   "86_Times_STEP_MAX_TIME_STP_540" : Time = PLC "86_Times".STEP_MAX_TIME_STP_540, 1 s
   "86_Times_STEP_MAX_TIME_STP_550" : Time = PLC "86_Times".STEP_MAX_TIME_STP_550, 1 s
   "86_Times_STEP_MAX_TIME_STP_560" : Time = PLC "86_Times".STEP_MAX_TIME_STP_560, 1 s
   "86_Times_STEP_MAX_TIME_STP_570" : Time = PLC "86_Times".STEP_MAX_TIME_STP_570, 1 s
   "86_Times_STEP_MAX_TIME_STP_580" : Time = PLC "86_Times".STEP_MAX_TIME_STP_580, 1 s
   "86_Times_STEP_MAX_TIME_STP_590" : Time = PLC "86_Times".STEP_MAX_TIME_STP_590, 1 s
   "86_Times_STEP_MAX_TIME_STP_600" : Time = PLC "86_Times".STEP_MAX_TIME_STP_600, 1 s
   "86_Times_STEP_MAX_TIME_STP_610" : Time = PLC "86_Times".STEP_MAX_TIME_STP_610, 1 s
   "86_Times_STEP_MAX_TIME_STP_620" : Time = PLC "86_Times".STEP_MAX_TIME_STP_620, 1 s
   "86_Times_STEP_MAX_TIME_STP_630" : Time = PLC "86_Times".STEP_MAX_TIME_STP_630, 1 s
   "150_GCU_LCL_CNTRL_DB_LCL_CNTRL_ACTV" : Bool = PLC "150_GCU_LCL_CNTRL_DB".LCL_CNTRL_ACTV, 1 s
   "150_GCU_LCL_CNTRL_DB_STRT_AIR" : Bool = PLC "150_GCU_LCL_CNTRL_DB".STRT_AIR, 1 s
   "150_GCU_LCL_CNTRL_DB_STRT_IG" : Bool = PLC "150_GCU_LCL_CNTRL_DB".STRT_IG, 1 s
   "150_GCU_LCL_CNTRL_DB_STOP" : Bool = PLC "150_GCU_LCL_CNTRL_DB".STOP, 1 s
   "150_GCU_LCL_CNTRL_DB_SYS_OK_FOR_LCL" : Bool = PLC "150_GCU_LCL_CNTRL_DB".SYS_OK_FOR_LCL, 1 s
   "150_GCU_LCL_CNTRL_DB_RUN_WITH_AIR" : Bool = PLC "150_GCU_LCL_CNTRL_DB".RUN_WITH_AIR, 1 s
   "150_GCU_LCL_CNTRL_DB_RUN_WITH_IG" : Bool = PLC "150_GCU_LCL_CNTRL_DB".RUN_WITH_IG, 1 s
   "80_From_HMI_Request_Auto" : Bool = PLC "80_From_HMI".Request_Auto, 1 s
   "80_From_HMI_Request_Manual" : Bool = PLC "80_From_HMI".Request_Manual, 1 s
   "80_From_HMI_RST_AUT_SEQ" : Bool = PLC "80_From_HMI".RST_AUT_SEQ, 1 s
   "141_P303_HRS_RUN_DB_HRS" : Int = PLC "141_P303_HRS_RUN_DB".HRS, 1 s
   "141_P303_HRS_RUN_DB_MINS" : Int = PLC "141_P303_HRS_RUN_DB".MINS, 1 s
   "141_P303_HRS_RUN_DB_SECS" : Int = PLC "141_P303_HRS_RUN_DB".SECS, 1 s
   "141_P303_HRS_RUN_DB_RST" : Bool = PLC "141_P303_HRS_RUN_DB".RST, 1 s
   "141_P303_HRS_RUN_DB_SRV_HRS" : Int = PLC "141_P303_HRS_RUN_DB".SRV_HRS, 1 s
   "141_P303_HRS_RUN_DB_SHRS_IP" : Int = PLC "141_P303_HRS_RUN_DB".SHRS_IP, 1 s
   "141_P303_HRS_RUN_DB_SRVC" : Bool = PLC "141_P303_HRS_RUN_DB".SRVC, 1 s
   "14_DQ_DATA_P_303" : Bool = PLC "14_DQ_DATA".P_303, 1 s
   "142_P304_HRS_RUN_DB_HRS" : Int = PLC "142_P304_HRS_RUN_DB".HRS, 1 s
   "142_P304_HRS_RUN_DB_MINS" : Int = PLC "142_P304_HRS_RUN_DB".MINS, 1 s
   "142_P304_HRS_RUN_DB_SECS" : Int = PLC "142_P304_HRS_RUN_DB".SECS, 1 s
   "142_P304_HRS_RUN_DB_RST" : Bool = PLC "142_P304_HRS_RUN_DB".RST, 1 s
   "142_P304_HRS_RUN_DB_SRV_HRS" : Int = PLC "142_P304_HRS_RUN_DB".SRV_HRS, 1 s
   "142_P304_HRS_RUN_DB_SHRS_IP" : Int = PLC "142_P304_HRS_RUN_DB".SHRS_IP, 1 s
   "142_P304_HRS_RUN_DB_SRVC" : Bool = PLC "142_P304_HRS_RUN_DB".SRVC, 1 s
   "14_DQ_DATA_P_304" : Bool = PLC "14_DQ_DATA".P_304, 1 s
   "100_GCU_AUTO_SEQ_DB_CRNT_STEP" : Int = PLC "100_GCU_AUTO_SEQ_DB".CRNT_STEP, 1 s
   "14_DQ_DATA_CV_422_APT" : Bool = PLC "14_DQ_DATA".CV_422_APT, 1 s
   "14_DQ_DATA_CV_421_6S" : Bool = PLC "14_DQ_DATA".CV_421_6S, 1 s
   "14_DQ_DATA_CV_422_6P" : Bool = PLC "14_DQ_DATA".CV_422_6P, 1 s
   "14_DQ_DATA_CV_421_5S" : Bool = PLC "14_DQ_DATA".CV_421_5S, 1 s
   "14_DQ_DATA_CV_422_5P" : Bool = PLC "14_DQ_DATA".CV_422_5P, 1 s
   "14_DQ_DATA_CV_421_4S" : Bool = PLC "14_DQ_DATA".CV_421_4S, 1 s
   "14_DQ_DATA_CV_422_4P" : Bool = PLC "14_DQ_DATA".CV_422_4P, 1 s
   "14_DQ_DATA_R3_SPR_DQ_138_7" : Bool = PLC "14_DQ_DATA".R3_SPR_DQ_138_7, 1 s
   "14_DQ_DATA_CV_421_3S" : Bool = PLC "14_DQ_DATA".CV_421_3S, 1 s
   "14_DQ_DATA_CV_422_3P" : Bool = PLC "14_DQ_DATA".CV_422_3P, 1 s
   "14_DQ_DATA_CV_421_1S" : Bool = PLC "14_DQ_DATA".CV_421_1S, 1 s
   "14_DQ_DATA_CV_422_1P" : Bool = PLC "14_DQ_DATA".CV_422_1P, 1 s
   "14_DQ_DATA_CV_422_FPT" : Bool = PLC "14_DQ_DATA".CV_422_FPT, 1 s
   "14_DQ_DATA_E_400_STP" : Bool = PLC "14_DQ_DATA".E_400_STP, 1 s
   "14_DQ_DATA_13P5" : Bool = PLC "14_DQ_DATA".13P5, 1 s
   "14_DQ_DATA_13P4" : Bool = PLC "14_DQ_DATA".13P4, 1 s
   "14_DQ_DATA_13P3" : Bool = PLC "14_DQ_DATA".13P3, 1 s
   "14_DQ_DATA_13P2" : Bool = PLC "14_DQ_DATA".13P2, 1 s
   "14_DQ_DATA_R3_SPR_DQ_139_7" : Bool = PLC "14_DQ_DATA".R3_SPR_DQ_139_7, 1 s
   "14_DQ_DATA_13P1" : Bool = PLC "14_DQ_DATA".13P1, 1 s
   "100_GCU_AUTO_SEQ_DB_RNG" : Bool = PLC "100_GCU_AUTO_SEQ_DB".RNG, 1 s

discrete alarms
   129: 'PIT-359 - HIGH HIGH', class IGG Alarms, trigger "60_Alarm_Data_IGG_ALARM_WORD_02" bit 1
   130: 'PIT-316 - HIGH HIGH', class IGG Alarms, trigger "60_Alarm_Data_IGG_ALARM_WORD_02" bit 3
   131: 'PIT-359 - LOW LOW', class IGG Alarms, trigger "60_Alarm_Data_IGG_ALARM_WORD_02" bit 0
   132: 'PIT-316 - LOW LOW', class IGG Alarms, trigger "60_Alarm_Data_IGG_ALARM_WORD_02" bit 2
   279: 'IGG_MESSAGE_WORD_02_BIT_14', class IGG Messages, trigger "64_Message_Data_IGG_MESSAGE_WORD_02" bit 6
   133: 'PIT-359 - HIGH HIGH', class IGG Alarms, trigger "60_Alarm_Data_IGG_ALARM_WORD_02" bit 4
   134: 'TIT-401 - HIGH HIGH', class IGG Alarms, trigger "60_Alarm_Data_IGG_ALARM_WORD_02" bit 10
   135: 'PIT-102 CA PRESSURE - FAULT', class IGG Alarms, trigger "60_Alarm_Data_IGG_ALARM_WORD_02" bit 9
   136: 'PIT-402 IG OUTLET PRESSURE - HIGH HIGH', class IGG Alarms, trigger "60_Alarm_Data_IGG_ALARM_WORD_02" bit 12
   137: 'PIT-402 IG OUTLET PRESSURE - LOW LOW', class IGG Alarms, trigger "60_Alarm_Data_IGG_ALARM_WORD_02" bit 11
   138: 'IGG_ALARM_WORD_02_BIT_14', class IGG Alarms, trigger "60_Alarm_Data_IGG_ALARM_WORD_02" bit 6
   139: 'IGG_ALARM_WORD_02_BIT_13', class IGG Alarms, trigger "60_Alarm_Data_IGG_ALARM_WORD_02" bit 5
   140: 'PIT-102 CA PRESSURE - LOW LOW', class IGG Alarms, trigger "60_Alarm_Data_IGG_ALARM_WORD_02" bit 8
   141: 'IGG_ALARM_WORD_02_BIT_15', class IGG Alarms, trigger "60_Alarm_Data_IGG_ALARM_WORD_02" bit 7
   142: 'EMERGENCY STOP ACTIVE', class IGG Alarms, trigger "60_Alarm_Data_IGG_ALARM_WORD_01" bit 15
   143: 'ATMOSPHERIC O2 SENSOR 1 - LOW LOW', class IGG Alarms, trigger "60_Alarm_Data_IGG_ALARM_WORD_01" bit 1
   144: 'BC ALARM ACTIVE', class IGG Alarms, trigger "60_Alarm_Data_IGG_ALARM_WORD_01" bit 0
   145: 'ATMOSPHERIC O2 SENSOR 2 - LOW LOW', class IGG Alarms, trigger "60_Alarm_Data_IGG_ALARM_WORD_01" bit 2
   146: 'E-500B FUEL PUMP - NOT RUNNING', class IGG Alarms, trigger "60_Alarm_Data_IGG_ALARM_WORD_01" bit 4
   147: 'E-500A FUEL PUMP - NOT RUNNING', class IGG Alarms, trigger "60_Alarm_Data_IGG_ALARM_WORD_01" bit 3
   383: 'BC_EVENT_WORD_02_BIT_6', class BC Events, trigger "66_Event_Data_BC_EVENT_WORD_02" bit 14
   382: 'BC_EVENT_WORD_02_BIT_5', class BC Events, trigger "66_Event_Data_BC_EVENT_WORD_02" bit 13
   384: 'BC_EVENT_WORD_02_BIT_7', class BC Events, trigger "66_Event_Data_BC_EVENT_WORD_02" bit 15
   278: 'IGG_MESSAGE_WORD_02_BIT_13', class IGG Messages, trigger "64_Message_Data_IGG_MESSAGE_WORD_02" bit 5
   277: 'IGG_MESSAGE_WORD_02_BIT_12', class IGG Messages, trigger "64_Message_Data_IGG_MESSAGE_WORD_02" bit 4
   148: 'P-301 CSW PUMP - TRIPPED', class IGG Alarms, trigger "60_Alarm_Data_IGG_ALARM_WORD_01" bit 11
   149: 'IGG AUTO INTERLOCKS NOT OK', class IGG Alarms, trigger "60_Alarm_Data_IGG_ALARM_WORD_01" bit 10
   150: 'E-500A FUEL PUMP - TRIPPED', class IGG Alarms, trigger "60_Alarm_Data_IGG_ALARM_WORD_01" bit 12
   151: 'E-139 CAB INVERTER - FAULT', class IGG Alarms, trigger "60_Alarm_Data_IGG_ALARM_WORD_01" bit 14
   152: 'E-500B FUEL PUMP - TRIPPED', class IGG Alarms, trigger "60_Alarm_Data_IGG_ALARM_WORD_01" bit 13
   153: 'IGG_ALARM_WORD_01_BIT_14', class IGG Alarms, trigger "60_Alarm_Data_IGG_ALARM_WORD_01" bit 6
   154: 'E-139 CAB NOT READY3', class IGG Alarms, trigger "60_Alarm_Data_IGG_ALARM_WORD_01" bit 5
   155: 'IGG_ALARM_WORD_01_BIT_15', class IGG Alarms, trigger "60_Alarm_Data_IGG_ALARM_WORD_01" bit 7
   156: 'SLAVE PLC HEART BEAT MISSING', class IGG Alarms, trigger "60_Alarm_Data_IGG_ALARM_WORD_01" bit 9
   157: 'MASTER PLC HEART BEAT MISSING', class IGG Alarms, trigger "60_Alarm_Data_IGG_ALARM_WORD_01" bit 8
   158: 'PIT-402 IG PRESSURE - OUT OF RANGE', class IGG Alarms, trigger "60_Alarm_Data_IGG_ALARM_WORD_02" bit 13
   55: 'IGG_ALARM_WORD_04_BIT_14', class IGG Alarms, trigger "60_Alarm_Data_IGG_ALARM_WORD_04" bit 6
   54: 'CORRECT PHASE ROTATION - FAULT', class IGG Alarms, trigger "60_Alarm_Data_IGG_ALARM_WORD_04" bit 5
   56: 'IGG_ALARM_WORD_04_BIT_15', class IGG Alarms, trigger "60_Alarm_Data_IGG_ALARM_WORD_04" bit 7
   58: 'CV-312 - FAULT', class IGG Alarms, trigger "60_Alarm_Data_IGG_ALARM_WORD_04" bit 9
   57: 'CV-311 - FAULT', class IGG Alarms, trigger "60_Alarm_Data_IGG_ALARM_WORD_04" bit 8
   50: 'TIT-319 INLET CSW TEMP - FAULT AND TIT-401 AND TIT-360 - FAULT', class IGG Alarms, trigger "60_Alarm_Data_IGG_ALARM_WORD_04" bit 1
   49: 'TIT-319 INLET CSW TEMP - FAULT AND TS-006 - FAULT', class IGG Alarms, trigger "60_Alarm_Data_IGG_ALARM_WORD_04" bit 0
   51: 'TIT-360 OUTLET CSW TEMP - HIGH HIGH0', class IGG Alarms, trigger "60_Alarm_Data_IGG_ALARM_WORD_04" bit 2
   53: 'E-139 NOT RUNNING2', class IGG Alarms, trigger "60_Alarm_Data_IGG_ALARM_WORD_04" bit 4
   52: 'TIT-360 OUTLET CSW TEMP - HIGH HIGH AND TIT-401 - FAULT', class IGG Alarms, trigger "60_Alarm_Data_IGG_ALARM_WORD_04" bit 3
   59: 'CV-321 - FAULT', class IGG Alarms, trigger "60_Alarm_Data_IGG_ALARM_WORD_04" bit 10
   65: 'IGG ALARM ACTIVE', class BC Alarms, trigger "60_Alarm_Data_BC_ALARM_WORD_01" bit 0
   282: 'IGG_MESSAGE_WORD_02_BIT_1', class IGG Messages, trigger "64_Message_Data_IGG_MESSAGE_WORD_02" bit 9
   66: 'PS-101 PRESSURE NOT PRESENT - FAULT', class BC Alarms, trigger "60_Alarm_Data_BC_ALARM_WORD_01" bit 1
   69: 'FD-001 FLAME SIGNAL - OUT OF RANGE', class BC Alarms, trigger "60_Alarm_Data_BC_ALARM_WORD_01" bit 4
   68: 'O2 SYSTEM POWER NOT HEALTHY', class BC Alarms, trigger "60_Alarm_Data_BC_ALARM_WORD_01" bit 3
   61: 'CV-401 - FAULT', class IGG Alarms, trigger "60_Alarm_Data_IGG_ALARM_WORD_04" bit 12
   60: 'CV-322 - FAULT', class IGG Alarms, trigger "60_Alarm_Data_IGG_ALARM_WORD_04" bit 11
   62: 'CV-431 - FAULT', class IGG Alarms, trigger "60_Alarm_Data_IGG_ALARM_WORD_04" bit 13
   64: 'SAFETY SYSTEM INTERLOCK', class IGG Alarms, trigger "60_Alarm_Data_IGG_ALARM_WORD_04" bit 15
   63: 'CV-432 - FAULT', class IGG Alarms, trigger "60_Alarm_Data_IGG_ALARM_WORD_04" bit 14
   35: 'TIT-315 SHELL CSW TEMP - HIGH HIGH AND TIT-401 - FAULT', class IGG Alarms, trigger "60_Alarm_Data_IGG_ALARM_WORD_03" bit 2
   34: 'TIT-315 SHELL CSW TEMP - HIGH HIGH AND TS-006 - FAULT', class IGG Alarms, trigger "60_Alarm_Data_IGG_ALARM_WORD_03" bit 1
   36: 'PIT-316 OUTLET CSW PRESSURE AND FS-317 - FAULT', class IGG Alarms, trigger "60_Alarm_Data_IGG_ALARM_WORD_03" bit 3
   38: 'PIT-316 OUTLET CSW PRESSURE AND TS-006 - FAULT', class IGG Alarms, trigger "60_Alarm_Data_IGG_ALARM_WORD_03" bit 5
   37: 'PIT-316 OUTLET CSW PRESSURE AND TIT-315 - FAULT', class IGG Alarms, trigger "60_Alarm_Data_IGG_ALARM_WORD_03" bit 4
   159: 'TIT-360 - HIGH HIGH', class IGG Alarms, trigger "60_Alarm_Data_IGG_ALARM_WORD_02" bit 15
   160: 'TIT-319 - HIGH HIGH', class IGG Alarms, trigger "60_Alarm_Data_IGG_ALARM_WORD_02" bit 14
   280: 'IGG_MESSAGE_WORD_02_BIT_15', class IGG Messages, trigger "64_Message_Data_IGG_MESSAGE_WORD_02" bit 7
   33: 'TIT-315 SHELL CSW TEMP - HIGH HIGH AND FS-317 - FAULT', class IGG Alarms, trigger "60_Alarm_Data_IGG_ALARM_WORD_03" bit 0
   70: 'E-600 O2 ANALYSER CONTENT - OUT OF RANGE', class BC Alarms, trigger "60_Alarm_Data_BC_ALARM_WORD_01" bit 5
   39: 'IGG_ALARM_WORD_03_BIT_14', class IGG Alarms, trigger "60_Alarm_Data_IGG_ALARM_WORD_03" bit 6
   46: 'TIT-401 IG TEMP - HIGH HIGH AND TIT-360 - FAULT', class IGG Alarms, trigger "60_Alarm_Data_IGG_ALARM_WORD_03" bit 13
   45: 'TIT-401 IG TEMP - HIGH HIGH AND TS-403 - FAULT', class IGG Alarms, trigger "60_Alarm_Data_IGG_ALARM_WORD_03" bit 12
   47: 'IGG_ALARM_WORD_03_BIT_6', class IGG Alarms, trigger "60_Alarm_Data_IGG_ALARM_WORD_03" bit 14
   281: 'IGG_MESSAGE_WORD_02_BIT_0', class IGG Messages, trigger "64_Message_Data_IGG_MESSAGE_WORD_02" bit 8
   48: 'IGG_ALARM_WORD_03_BIT_7', class IGG Alarms, trigger "60_Alarm_Data_IGG_ALARM_WORD_03" bit 15
   41: 'PIT-112/113 TIER ALARM - PRESSURE NOT OK', class IGG Alarms, trigger "60_Alarm_Data_IGG_ALARM_WORD_03" bit 8
   40: 'IGG_ALARM_WORD_03_BIT_15', class IGG Alarms, trigger "60_Alarm_Data_IGG_ALARM_WORD_03" bit 7
   42: 'PIT-102 CA PRESSURE - LOW LOW AND FDU - FAULT', class IGG Alarms, trigger "60_Alarm_Data_IGG_ALARM_WORD_03" bit 9
   44: 'IGG ALARM WORD', class IGG Alarms, trigger "60_Alarm_Data_IGG_ALARM_WORD_03" bit 11
   43: 'PIT-102 CA PRESSURE - LOW LOW AND PIT-402 - FAULT', class IGG Alarms, trigger "60_Alarm_Data_IGG_ALARM_WORD_03" bit 10
   381: 'BC_EVENT_WORD_02_BIT_4', class BC Events, trigger "66_Event_Data_BC_EVENT_WORD_02" bit 12
   330: 'IGG_EVENT_WORD_01_BIT_1', class IGG Events, trigger "66_Event_Data_IGG_EVENT_WORD_01" bit 9
   329: 'IGG_EVENT_WORD_01_BIT_0', class IGG Events, trigger "66_Event_Data_IGG_EVENT_WORD_01" bit 8
   331: 'IGG_EVENT_WORD_01_BIT_2', class IGG Events, trigger "66_Event_Data_IGG_EVENT_WORD_01" bit 10
   333: 'IGG_EVENT_WORD_01_BIT_4', class IGG Events, trigger "66_Event_Data_IGG_EVENT_WORD_01" bit 12
   332: 'IGG_EVENT_WORD_01_BIT_3', class IGG Events, trigger "66_Event_Data_IGG_EVENT_WORD_01" bit 11
   325: 'IGG_EVENT_WORD_01_BIT_12', class IGG Events, trigger "66_Event_Data_IGG_EVENT_WORD_01" bit 4
   324: 'IGG_EVENT_WORD_01_BIT_11', class IGG Events, trigger "66_Event_Data_IGG_EVENT_WORD_01" bit 3
   326: 'IGG_EVENT_WORD_01_BIT_13', class IGG Events, trigger "66_Event_Data_IGG_EVENT_WORD_01" bit 5
   328: 'IGG_EVENT_WORD_01_BIT_15', class IGG Events, trigger "66_Event_Data_IGG_EVENT_WORD_01" bit 7
   327: 'IGG_EVENT_WORD_01_BIT_14', class IGG Events, trigger "66_Event_Data_IGG_EVENT_WORD_01" bit 6
   338: 'IGG_EVENT_WORD_02_BIT_9', class IGG Events, trigger "66_Event_Data_IGG_EVENT_WORD_02" bit 1
   337: 'IGG_EVENT_WORD_02_BIT_8', class IGG Events, trigger "66_Event_Data_IGG_EVENT_WORD_02" bit 0
   339: 'IGG_EVENT_WORD_02_BIT_10', class IGG Events, trigger "66_Event_Data_IGG_EVENT_WORD_02" bit 2
   341: 'IGG_EVENT_WORD_02_BIT_12', class IGG Events, trigger "66_Event_Data_IGG_EVENT_WORD_02" bit 4
   340: 'IGG_EVENT_WORD_02_BIT_11', class IGG Events, trigger "66_Event_Data_IGG_EVENT_WORD_02" bit 3
   335: 'IGG_EVENT_WORD_01_BIT_6', class IGG Events, trigger "66_Event_Data_IGG_EVENT_WORD_01" bit 14
   334: 'IGG_EVENT_WORD_01_BIT_5', class IGG Events, trigger "66_Event_Data_IGG_EVENT_WORD_01" bit 13
   336: 'IGG_EVENT_WORD_01_BIT_7', class IGG Events, trigger "66_Event_Data_IGG_EVENT_WORD_01" bit 15
   276: 'IGG_MESSAGE_WORD_02_BIT_11', class IGG Messages, trigger "64_Message_Data_IGG_MESSAGE_WORD_02" bit 3
   259: 'IGG_MESSAGE_WORD_01_BIT_10', class IGG Messages, trigger "64_Message_Data_IGG_MESSAGE_WORD_01" bit 2
   267: 'IGG_MESSAGE_WORD_01_BIT_2', class IGG Messages, trigger "64_Message_Data_IGG_MESSAGE_WORD_01" bit 10
   268: 'IGG_MESSAGE_WORD_01_BIT_3', class IGG Messages, trigger "64_Message_Data_IGG_MESSAGE_WORD_01" bit 11
   273: 'IGG_MESSAGE_WORD_02_BIT_8', class IGG Messages, trigger "64_Message_Data_IGG_MESSAGE_WORD_02" bit 0
   265: 'IGG_MESSAGE_WORD_01_BIT_0', class IGG Messages, trigger "64_Message_Data_IGG_MESSAGE_WORD_01" bit 8
   266: 'IGG_MESSAGE_WORD_01_BIT_1', class IGG Messages, trigger "64_Message_Data_IGG_MESSAGE_WORD_01" bit 9
   272: 'IGG_MESSAGE_WORD_01_BIT_7', class IGG Messages, trigger "64_Message_Data_IGG_MESSAGE_WORD_01" bit 15
   67: 'E-600 O2 ANALYSER SYSTEM - FAIL', class BC Alarms, trigger "60_Alarm_Data_BC_ALARM_WORD_01" bit 2
   271: 'IGG_MESSAGE_WORD_01_BIT_6', class IGG Messages, trigger "64_Message_Data_IGG_MESSAGE_WORD_01" bit 14
   269: 'IGG_MESSAGE_WORD_01_BIT_4', class IGG Messages, trigger "64_Message_Data_IGG_MESSAGE_WORD_01" bit 12
   270: 'IGG_MESSAGE_WORD_01_BIT_5', class IGG Messages, trigger "64_Message_Data_IGG_MESSAGE_WORD_01" bit 13
   260: 'IGG_MESSAGE_WORD_01_BIT_11', class IGG Messages, trigger "64_Message_Data_IGG_MESSAGE_WORD_01" bit 3
   275: 'IGG_MESSAGE_WORD_02_BIT_10', class IGG Messages, trigger "64_Message_Data_IGG_MESSAGE_WORD_02" bit 2
   321: 'IGG_EVENT_WORD_01_BIT_8', class IGG Events, trigger "66_Event_Data_IGG_EVENT_WORD_01" bit 0
   323: 'IGG_EVENT_WORD_01_BIT_10', class IGG Events, trigger "66_Event_Data_IGG_EVENT_WORD_01" bit 2
   322: 'IGG_EVENT_WORD_01_BIT_9', class IGG Events, trigger "66_Event_Data_IGG_EVENT_WORD_01" bit 1
   264: 'IGG_MESSAGE_WORD_01_BIT_15', class IGG Messages, trigger "64_Message_Data_IGG_MESSAGE_WORD_01" bit 7
   274: 'IGG_MESSAGE_WORD_02_BIT_9', class IGG Messages, trigger "64_Message_Data_IGG_MESSAGE_WORD_02" bit 1
   263: 'IGG_MESSAGE_WORD_01_BIT_14', class IGG Messages, trigger "64_Message_Data_IGG_MESSAGE_WORD_01" bit 6
   261: 'IGG_MESSAGE_WORD_01_BIT_12', class IGG Messages, trigger "64_Message_Data_IGG_MESSAGE_WORD_01" bit 4
   262: 'IGG_MESSAGE_WORD_01_BIT_13', class IGG Messages, trigger "64_Message_Data_IGG_MESSAGE_WORD_01" bit 5
   342: 'IGG_EVENT_WORD_02_BIT_13', class IGG Events, trigger "66_Event_Data_IGG_EVENT_WORD_02" bit 5
   367: 'BC_EVENT_WORD_01_BIT_6', class BC Events, trigger "66_Event_Data_BC_EVENT_WORD_01" bit 14
   366: 'BC_EVENT_WORD_01_BIT_5', class BC Events, trigger "66_Event_Data_BC_EVENT_WORD_01" bit 13
   368: 'BC_EVENT_WORD_01_BIT_7', class BC Events, trigger "66_Event_Data_BC_EVENT_WORD_01" bit 15
   370: 'BC_EVENT_WORD_02_BIT_9', class BC Events, trigger "66_Event_Data_BC_EVENT_WORD_02" bit 1
   369: 'BC_EVENT_WORD_02_BIT_8', class BC Events, trigger "66_Event_Data_BC_EVENT_WORD_02" bit 0
   362: 'BC_EVENT_WORD_01_BIT_1', class BC Events, trigger "66_Event_Data_BC_EVENT_WORD_01" bit 9
   361: 'BC_EVENT_WORD_01_BIT_0', class BC Events, trigger "66_Event_Data_BC_EVENT_WORD_01" bit 8
   363: 'BC_EVENT_WORD_01_BIT_2', class BC Events, trigger "66_Event_Data_BC_EVENT_WORD_01" bit 10
   365: 'BC_EVENT_WORD_01_BIT_4', class BC Events, trigger "66_Event_Data_BC_EVENT_WORD_01" bit 12
   364: 'BC_EVENT_WORD_01_BIT_3', class BC Events, trigger "66_Event_Data_BC_EVENT_WORD_01" bit 11
   377: 'BC_EVENT_WORD_02_BIT_0', class BC Events, trigger "66_Event_Data_BC_EVENT_WORD_02" bit 8
   376: 'BC_EVENT_WORD_02_BIT_15', class BC Events, trigger "66_Event_Data_BC_EVENT_WORD_02" bit 7
   378: 'BC_EVENT_WORD_02_BIT_1', class BC Events, trigger "66_Event_Data_BC_EVENT_WORD_02" bit 9
   380: 'BC_EVENT_WORD_02_BIT_3', class BC Events, trigger "66_Event_Data_BC_EVENT_WORD_02" bit 11
   379: 'BC_EVENT_WORD_02_BIT_2', class BC Events, trigger "66_Event_Data_BC_EVENT_WORD_02" bit 10
   372: 'BC_EVENT_WORD_02_BIT_11', class BC Events, trigger "66_Event_Data_BC_EVENT_WORD_02" bit 3
   371: 'BC_EVENT_WORD_02_BIT_10', class BC Events, trigger "66_Event_Data_BC_EVENT_WORD_02" bit 2
   373: 'BC_EVENT_WORD_02_BIT_12', class BC Events, trigger "66_Event_Data_BC_EVENT_WORD_02" bit 4
   375: 'BC_EVENT_WORD_02_BIT_14', class BC Events, trigger "66_Event_Data_BC_EVENT_WORD_02" bit 6
   374: 'BC_EVENT_WORD_02_BIT_13', class BC Events, trigger "66_Event_Data_BC_EVENT_WORD_02" bit 5
   349: 'IGG_EVENT_WORD_02_BIT_4', class IGG Events, trigger "66_Event_Data_IGG_EVENT_WORD_02" bit 12
   348: 'IGG_EVENT_WORD_02_BIT_3', class IGG Events, trigger "66_Event_Data_IGG_EVENT_WORD_02" bit 11
   350: 'IGG_EVENT_WORD_02_BIT_5', class IGG Events, trigger "66_Event_Data_IGG_EVENT_WORD_02" bit 13
   352: 'IGG_EVENT_WORD_02_BIT_7', class IGG Events, trigger "66_Event_Data_IGG_EVENT_WORD_02" bit 15
   351: 'IGG_EVENT_WORD_02_BIT_6', class IGG Events, trigger "66_Event_Data_IGG_EVENT_WORD_02" bit 14
   344: 'IGG_EVENT_WORD_02_BIT_15', class IGG Events, trigger "66_Event_Data_IGG_EVENT_WORD_02" bit 7
   343: 'IGG_EVENT_WORD_02_BIT_14', class IGG Events, trigger "66_Event_Data_IGG_EVENT_WORD_02" bit 6
   345: 'IGG_EVENT_WORD_02_BIT_0', class IGG Events, trigger "66_Event_Data_IGG_EVENT_WORD_02" bit 8
   347: 'IGG_EVENT_WORD_02_BIT_2', class IGG Events, trigger "66_Event_Data_IGG_EVENT_WORD_02" bit 10
   346: 'IGG_EVENT_WORD_02_BIT_1', class IGG Events, trigger "66_Event_Data_IGG_EVENT_WORD_02" bit 9
   357: 'BC_EVENT_WORD_01_BIT_12', class BC Events, trigger "66_Event_Data_BC_EVENT_WORD_01" bit 4
   356: 'BC_EVENT_WORD_01_BIT_11', class BC Events, trigger "66_Event_Data_BC_EVENT_WORD_01" bit 3
   358: 'BC_EVENT_WORD_01_BIT_13', class BC Events, trigger "66_Event_Data_BC_EVENT_WORD_01" bit 5
   360: 'BC_EVENT_WORD_01_BIT_15', class BC Events, trigger "66_Event_Data_BC_EVENT_WORD_01" bit 7
   359: 'BC_EVENT_WORD_01_BIT_14', class BC Events, trigger "66_Event_Data_BC_EVENT_WORD_01" bit 6
   257: 'IGG_MESSAGE_WORD_01_BIT_8', class IGG Messages, trigger "64_Message_Data_IGG_MESSAGE_WORD_01" bit 0
   258: 'IGG_MESSAGE_WORD_01_BIT_9', class IGG Messages, trigger "64_Message_Data_IGG_MESSAGE_WORD_01" bit 1
   353: 'BC_EVENT_WORD_01_BIT_8', class BC Events, trigger "66_Event_Data_BC_EVENT_WORD_01" bit 0
   355: 'BC_EVENT_WORD_01_BIT_10', class BC Events, trigger "66_Event_Data_BC_EVENT_WORD_01" bit 2
   354: 'BC_EVENT_WORD_01_BIT_9', class BC Events, trigger "66_Event_Data_BC_EVENT_WORD_01" bit 1
   114: 'P-305 FRESH WATER PUMP - TRIPPED', class BC Alarms, trigger "60_Alarm_Data_BC_ALARM_WORD_04" bit 1
   113: 'LS-001 IGG QUENCH CHAMBER LEVEL - HIGH', class BC Alarms, trigger "60_Alarm_Data_BC_ALARM_WORD_04" bit 0
   116: 'BC_ALARM_WORD_04_BIT_11', class BC Alarms, trigger "60_Alarm_Data_BC_ALARM_WORD_04" bit 3
   115: 'BC_ALARM_WORD_04_BIT_10', class BC Alarms, trigger "60_Alarm_Data_BC_ALARM_WORD_04" bit 2
   284: 'IGG_MESSAGE_WORD_02_BIT_3', class IGG Messages, trigger "64_Message_Data_IGG_MESSAGE_WORD_02" bit 11
   112: 'BC_ALARM_WORD_3_BIT_15', class BC Alarms, trigger "60_Alarm_Data_BC_ALARM_WORD_03" bit 15
   315: 'BC_MESSAGE_WORD_02_BIT_2', class BC Messages, trigger "64_Message_Data_BC_MESSAGE_WORD_02" bit 10
   316: 'BC_MESSAGE_WORD_02_BIT_3', class BC Messages, trigger "64_Message_Data_BC_MESSAGE_WORD_02" bit 11
   122: 'TS-006 IG SHELL TEMP HI SWITCH AND TIT-360 - FAULT', class BC Alarms, trigger "60_Alarm_Data_BC_ALARM_WORD_04" bit 9
   121: 'TS-006 IGG SHELL TEMPERATURE - HIGH', class BC Alarms, trigger "60_Alarm_Data_BC_ALARM_WORD_04" bit 8
   124: 'TS-403 IG TEMP - HIGH HIGH SWITCH AND TIT-401 - FAULT', class BC Alarms, trigger "60_Alarm_Data_BC_ALARM_WORD_04" bit 11
   123: 'TS-006 IG SHELL TEMP HI SWITCH AND TIT-401 - FAULT', class BC Alarms, trigger "60_Alarm_Data_BC_ALARM_WORD_04" bit 10
   297: 'BC_MESSAGE_WORD_01_BIT_0', class BC Messages, trigger "64_Message_Data_BC_MESSAGE_WORD_01" bit 8
   117: 'BC_ALARM_WORD_04_BIT_12', class BC Alarms, trigger "60_Alarm_Data_BC_ALARM_WORD_04" bit 4
   120: 'BC_ALARM_WORD_04_BIT_15', class BC Alarms, trigger "60_Alarm_Data_BC_ALARM_WORD_04" bit 7
   119: 'BC_ALARM_WORD_04_BIT_14', class BC Alarms, trigger "60_Alarm_Data_BC_ALARM_WORD_04" bit 6
   111: 'BC_ALARM_WORD_03_BIT_6', class BC Alarms, trigger "60_Alarm_Data_BC_ALARM_WORD_03" bit 14
   100: 'FS-317 JACKET COOLING WATER FLOW SWITCH - FAULT AND FS-320 - FAULT AND PIT 360 - FAULT', class BC Alarms, trigger "60_Alarm_Data_BC_ALARM_WORD_03" bit 3
   99: 'FS-320 COOLING WATER FLOW SWITCH - FAULT AND TIT-401 - FAULT0', class BC Alarms, trigger "60_Alarm_Data_BC_ALARM_WORD_03" bit 2
   102: 'FS-317 JACKET COOLING WATER FLOW SWITCH - FAULT AND TIT-401 - FAULT', class BC Alarms, trigger "60_Alarm_Data_BC_ALARM_WORD_03" bit 5
   101: 'FS-317 JACKET COOLING WATER FLOW SWITCH FASULT AND TIT-360 - FAULT', class BC Alarms, trigger "60_Alarm_Data_BC_ALARM_WORD_03" bit 4
   317: 'BC_MESSAGE_WORD_02_BIT_4', class BC Messages, trigger "64_Message_Data_BC_MESSAGE_WORD_02" bit 12
   318: 'BC_MESSAGE_WORD_02_BIT_5', class BC Messages, trigger "64_Message_Data_BC_MESSAGE_WORD_02" bit 13
   98: 'FS-320 COOLING WATER FLOW SWITCH - FAULT AND TIT-360 - FAULT', class BC Alarms, trigger "60_Alarm_Data_BC_ALARM_WORD_03" bit 1
   97: 'FS-320 COOLING WATER FLOW SWITCH - FAULT AND FS-317 - FAULT', class BC Alarms, trigger "60_Alarm_Data_BC_ALARM_WORD_03" bit 0
   108: 'PIT-112 INSTRUMENT AIR PRESSURE - FAULT AND FS-115 - FAULT', class BC Alarms, trigger "60_Alarm_Data_BC_ALARM_WORD_03" bit 11
   107: 'PIT-112 INSTRUMENT AIR PRESSURE - FAULT', class BC Alarms, trigger "60_Alarm_Data_BC_ALARM_WORD_03" bit 10
   110: 'FS-115 MAIN BURNER ATOMISING AIR FLOW SWITCH - FAULT AND PIT-113 - FAULT', class BC Alarms, trigger "60_Alarm_Data_BC_ALARM_WORD_03" bit 13
   109: 'FS-115 MAIN BURNER ATOMISING AIR FLOW SWITCH - FAULT AND CV 114 CLOSE', class BC Alarms, trigger "60_Alarm_Data_BC_ALARM_WORD_03" bit 12
   104: 'TS-403 IG VENT TEMPERATURE HIGH', class BC Alarms, trigger "60_Alarm_Data_BC_ALARM_WORD_03" bit 7
   103: 'BC_ALARM_WORD_03_BIT_14', class BC Alarms, trigger "60_Alarm_Data_BC_ALARM_WORD_03" bit 6
   106: 'FS-123 PILOT BURNER AIR FLOW SWITCH - FAULT AND PIT-112 LOW LOW', class BC Alarms, trigger "60_Alarm_Data_BC_ALARM_WORD_03" bit 9
   105: 'FS-123 PILOT BURNER AIR FLOW SWITCH - FAULT AND PIT-112 HIGH HIGH', class BC Alarms, trigger "60_Alarm_Data_BC_ALARM_WORD_03" bit 8
   305: 'BC_MESSAGE_WORD_02_BIT_8', class BC Messages, trigger "64_Message_Data_BC_MESSAGE_WORD_02" bit 0
   306: 'BC_MESSAGE_WORD_02_BIT_9', class BC Messages, trigger "64_Message_Data_BC_MESSAGE_WORD_02" bit 1
   304: 'BC_MESSAGE_WORD_01_BIT_7', class BC Messages, trigger "64_Message_Data_BC_MESSAGE_WORD_01" bit 15
   294: 'BC_MESSAGE_WORD_01_BIT_13', class BC Messages, trigger "64_Message_Data_BC_MESSAGE_WORD_01" bit 5
   293: 'BC_MESSAGE_WORD_01_BIT_12', class BC Messages, trigger "64_Message_Data_BC_MESSAGE_WORD_01" bit 4
   309: 'BC_MESSAGE_WORD_02_BIT_12', class BC Messages, trigger "64_Message_Data_BC_MESSAGE_WORD_02" bit 4
   307: 'BC_MESSAGE_WORD_02_BIT_10', class BC Messages, trigger "64_Message_Data_BC_MESSAGE_WORD_02" bit 2
   308: 'BC_MESSAGE_WORD_02_BIT_11', class BC Messages, trigger "64_Message_Data_BC_MESSAGE_WORD_02" bit 3
   300: 'BC_MESSAGE_WORD_01_BIT_3', class BC Messages, trigger "64_Message_Data_BC_MESSAGE_WORD_01" bit 11
   296: 'BC_MESSAGE_WORD_01_BIT_15', class BC Messages, trigger "64_Message_Data_BC_MESSAGE_WORD_01" bit 7
   298: 'BC_MESSAGE_WORD_01_BIT_1', class BC Messages, trigger "64_Message_Data_BC_MESSAGE_WORD_01" bit 9
   299: 'BC_MESSAGE_WORD_01_BIT_2', class BC Messages, trigger "64_Message_Data_BC_MESSAGE_WORD_01" bit 10
   295: 'BC_MESSAGE_WORD_01_BIT_14', class BC Messages, trigger "64_Message_Data_BC_MESSAGE_WORD_01" bit 6
   303: 'BC_MESSAGE_WORD_01_BIT_6', class BC Messages, trigger "64_Message_Data_BC_MESSAGE_WORD_01" bit 14
   301: 'BC_MESSAGE_WORD_01_BIT_4', class BC Messages, trigger "64_Message_Data_BC_MESSAGE_WORD_01" bit 12
   302: 'BC_MESSAGE_WORD_01_BIT_5', class BC Messages, trigger "64_Message_Data_BC_MESSAGE_WORD_01" bit 13
   310: 'BC_MESSAGE_WORD_02_BIT_13', class BC Messages, trigger "64_Message_Data_BC_MESSAGE_WORD_02" bit 5
   285: 'IGG_MESSAGE_WORD_02_BIT_4', class IGG Messages, trigger "64_Message_Data_IGG_MESSAGE_WORD_02" bit 12
   314: 'BC_MESSAGE_WORD_02_BIT_1', class BC Messages, trigger "64_Message_Data_BC_MESSAGE_WORD_02" bit 9
   287: 'IGG_MESSAGE_WORD_02_BIT_6', class IGG Messages, trigger "64_Message_Data_IGG_MESSAGE_WORD_02" bit 14
   286: 'IGG_MESSAGE_WORD_02_BIT_5', class IGG Messages, trigger "64_Message_Data_IGG_MESSAGE_WORD_02" bit 13
   126: 'PIT-113 IGG MAIN ATOM AIR PRESSURE - FAULT', class BC Alarms, trigger "60_Alarm_Data_BC_ALARM_WORD_04" bit 13
   125: 'TS-403 IG TEMP - HIGH HIGH SWITCH AND TIT-360 - FAULT', class BC Alarms, trigger "60_Alarm_Data_BC_ALARM_WORD_04" bit 12
   128: 'TIT-202 IGG INLET FUEL TEMP', class BC Alarms, trigger "60_Alarm_Data_BC_ALARM_WORD_04" bit 15
   127: 'PIT-205 IGG MAIN FUEL PRESSURE - FAULT', class BC Alarms, trigger "60_Alarm_Data_BC_ALARM_WORD_04" bit 14
   313: 'BC_MESSAGE_WORD_02_BIT_0', class BC Messages, trigger "64_Message_Data_BC_MESSAGE_WORD_02" bit 8
   292: 'BC_MESSAGE_WORD_01_BIT_11', class BC Messages, trigger "64_Message_Data_BC_MESSAGE_WORD_01" bit 3
   311: 'BC_MESSAGE_WORD_02_BIT_14', class BC Messages, trigger "64_Message_Data_BC_MESSAGE_WORD_02" bit 6
   312: 'BC_MESSAGE_WORD_02_BIT_15', class BC Messages, trigger "64_Message_Data_BC_MESSAGE_WORD_02" bit 7
   289: 'BC_MESSAGE_WORD_01_BIT_8', class BC Messages, trigger "64_Message_Data_BC_MESSAGE_WORD_01" bit 0
   288: 'IGG_MESSAGE_WORD_02_BIT_7', class IGG Messages, trigger "64_Message_Data_IGG_MESSAGE_WORD_02" bit 15
   291: 'BC_MESSAGE_WORD_01_BIT_10', class BC Messages, trigger "64_Message_Data_BC_MESSAGE_WORD_01" bit 2
   290: 'BC_MESSAGE_WORD_01_BIT_9', class BC Messages, trigger "64_Message_Data_BC_MESSAGE_WORD_01" bit 1
   93: 'BC_ALARM_WORD_02_BIT_4', class BC Alarms, trigger "60_Alarm_Data_BC_ALARM_WORD_02" bit 12
   75: 'BC AUTO INTERLOCKS NOT OK', class BC Alarms, trigger "60_Alarm_Data_BC_ALARM_WORD_01" bit 10
   88: 'BC_ALARM_WORD_02_BIT_15', class BC Alarms, trigger "60_Alarm_Data_BC_ALARM_WORD_02" bit 7
   283: 'IGG_MESSAGE_WORD_02_BIT_2', class IGG Messages, trigger "64_Message_Data_IGG_MESSAGE_WORD_02" bit 10
   320: 'BC_MESSAGE_WORD_02_BIT_7', class BC Messages, trigger "64_Message_Data_BC_MESSAGE_WORD_02" bit 15
   94: 'BC_ALARM_WORD_02_BIT_5', class BC Alarms, trigger "60_Alarm_Data_BC_ALARM_WORD_02" bit 13
   74: 'IGNITER POWER NOT HEALTHY', class BC Alarms, trigger "60_Alarm_Data_BC_ALARM_WORD_01" bit 9
   79: 'PILOT FLAME PURGE SEQUENCE FAILURE', class BC Alarms, trigger "60_Alarm_Data_BC_ALARM_WORD_01" bit 14
   80: 'FD-001 FLAME DETECTION UNIT NOT HEALTHY', class BC Alarms, trigger "60_Alarm_Data_BC_ALARM_WORD_01" bit 15
   84: 'PIT-204 FUEL OIL INLET PRESSURE LOW LOW AND PIT-205 - FAULT', class BC Alarms, trigger "60_Alarm_Data_BC_ALARM_WORD_02" bit 3
   90: 'NO FLOW AT FS-320', class BC Alarms, trigger "60_Alarm_Data_BC_ALARM_WORD_02" bit 9
   91: 'BC_ALARM_WORD_02_BIT_2', class BC Alarms, trigger "60_Alarm_Data_BC_ALARM_WORD_02" bit 10
   83: 'BC_ALARM_WORD_02_BIT_10', class BC Alarms, trigger "60_Alarm_Data_BC_ALARM_WORD_02" bit 2
   82: 'PIT-204 FUEL OIL INLET PRESSURE READING - FAULT AND CV-206 AND CV-207 - CLOSED', class BC Alarms, trigger "60_Alarm_Data_BC_ALARM_WORD_02" bit 1
   76: 'FDU POWER NOT HEALTHY', class BC Alarms, trigger "60_Alarm_Data_BC_ALARM_WORD_01" bit 11
   89: 'NO FLOW AT FS-317', class BC Alarms, trigger "60_Alarm_Data_BC_ALARM_WORD_02" bit 8
   95: 'BC_ALARM_WORD_02_BIT_6', class BC Alarms, trigger "60_Alarm_Data_BC_ALARM_WORD_02" bit 14
   87: 'PIT-204 FUEL OIL INLET PRESSURE - HIGH HIGH AND CV-206 AND CV-207 CLOSED', class BC Alarms, trigger "60_Alarm_Data_BC_ALARM_WORD_02" bit 6
   85: 'PIT-204 FUEL OIL INLET PRESSURE - LOW LOW', class BC Alarms, trigger "60_Alarm_Data_BC_ALARM_WORD_02" bit 4
   71: 'E-600 O2 ANALYSER CONTENT - LOW LOW', class BC Alarms, trigger "60_Alarm_Data_BC_ALARM_WORD_01" bit 6
   77: 'PILOT FLAME IGNITION SEQUENCE FAILURE', class BC Alarms, trigger "60_Alarm_Data_BC_ALARM_WORD_01" bit 12
   86: 'PIT-204 FUEL OIL INLET PRESSURE - HIGH HIGH AND PIT-205 - FAULT', class BC Alarms, trigger "60_Alarm_Data_BC_ALARM_WORD_02" bit 5
   78: 'MAIN BURNER FLAME SEQUENCE FAILURE', class BC Alarms, trigger "60_Alarm_Data_BC_ALARM_WORD_01" bit 13
   92: 'BC_ALARM_WORD_02_BIT_3', class BC Alarms, trigger "60_Alarm_Data_BC_ALARM_WORD_02" bit 11
   96: 'BC_ALARM_WORD_02_BIT_7', class BC Alarms, trigger "60_Alarm_Data_BC_ALARM_WORD_02" bit 15
   118: 'BC_ALARM_WORD_04_BIT_13', class BC Alarms, trigger "60_Alarm_Data_BC_ALARM_WORD_04" bit 5
   72: 'E-600 O2 ANALYSER CONTENT - HIGH HIGH', class BC Alarms, trigger "60_Alarm_Data_BC_ALARM_WORD_01" bit 7
   73: 'MASTER PLC HEART BEAT MISSING', class BC Alarms, trigger "60_Alarm_Data_BC_ALARM_WORD_01" bit 8
   81: 'PIT-204 FUEL OIL INLET PRESSURE READING - FAULT AND PIT-205 - FAULT', class BC Alarms, trigger "60_Alarm_Data_BC_ALARM_WORD_02" bit 0
   319: 'BC_MESSAGE_WORD_02_BIT_6', class BC Messages, trigger "64_Message_Data_BC_MESSAGE_WORD_02" bit 14
   385: 'IGG_WARNING_WORD_01_BIT_8', class IGG Warnings, trigger "62_Warning_Data_IGG_WARNING_WORD_01" bit 0
   386: 'IGG_WARNING_WORD_01_BIT_9', class IGG Warnings, trigger "62_Warning_Data_IGG_WARNING_WORD_01" bit 1
   387: 'IGG_WARNING_WORD_01_BIT_10', class IGG Warnings, trigger "62_Warning_Data_IGG_WARNING_WORD_01" bit 2
   388: 'IGG_WARNING_WORD_01_BIT_11', class IGG Warnings, trigger "62_Warning_Data_IGG_WARNING_WORD_01" bit 3
   389: 'IGG_WARNING_WORD_01_BIT_12', class IGG Warnings, trigger "62_Warning_Data_IGG_WARNING_WORD_01" bit 4
   390: 'IGG_WARNING_WORD_01_BIT_13', class IGG Warnings, trigger "62_Warning_Data_IGG_WARNING_WORD_01" bit 5
   391: 'IGG_WARNING_WORD_01_BIT_14', class IGG Warnings, trigger "62_Warning_Data_IGG_WARNING_WORD_01" bit 6
   392: 'IGG_WARNING_WORD_01_BIT_15', class IGG Warnings, trigger "62_Warning_Data_IGG_WARNING_WORD_01" bit 7
   393: '31B1 ATMOSPHERIC O2 SENSOR - LOW', class IGG Warnings, trigger "62_Warning_Data_IGG_WARNING_WORD_01" bit 8
   394: '31B2 ATMOSPHERIC O2 SENSOR - LOW', class IGG Warnings, trigger "62_Warning_Data_IGG_WARNING_WORD_01" bit 9
   395: '31B1 ATMOSPHERIC O2 SENSOR - LOW LOW', class IGG Warnings, trigger "62_Warning_Data_IGG_WARNING_WORD_01" bit 10
   396: '31B2 ATMOSPHERIC O2 SENSOR - LOW LOW', class IGG Warnings, trigger "62_Warning_Data_IGG_WARNING_WORD_01" bit 11
   397: 'IGG_WARNING_WORD_01_BIT_4', class IGG Warnings, trigger "62_Warning_Data_IGG_WARNING_WORD_01" bit 12